(* Logix 5000 project; controller PLC_MCC1300_75F1 vendor 1 type 14 code 166 rev 32.11; software revision 32.04; part 13 of 83 *)
(* tags used below, declared in another part *)
   M302SpeedUp : MAC_SpeedUp;
   TMP_d : DINT;
   TMP_xPositioning : BOOL;
   TMP_xReverse : BOOL;
   TMP_xRun : BOOL;
   xAlwaysOFF : BOOL;
   Z300_Conveyor : UDT_StandConv[29];
   Z300_Conveyor_Conf : UDT_Conveyor_Config[29];
   Z300_Conveyor_HMW : MAC_Conveyor_ZC_HMW[29];
   Z300_Conveyor_IN_MOTION : MAC_Conveyor_ZC_IN_MOTION[29];
   Z301_HMR : MAC_Zone_ML_HMR;
(* CommandLogic, continued *)

ROUTINE M302M5_Conveyor_Output   (* ladder *)
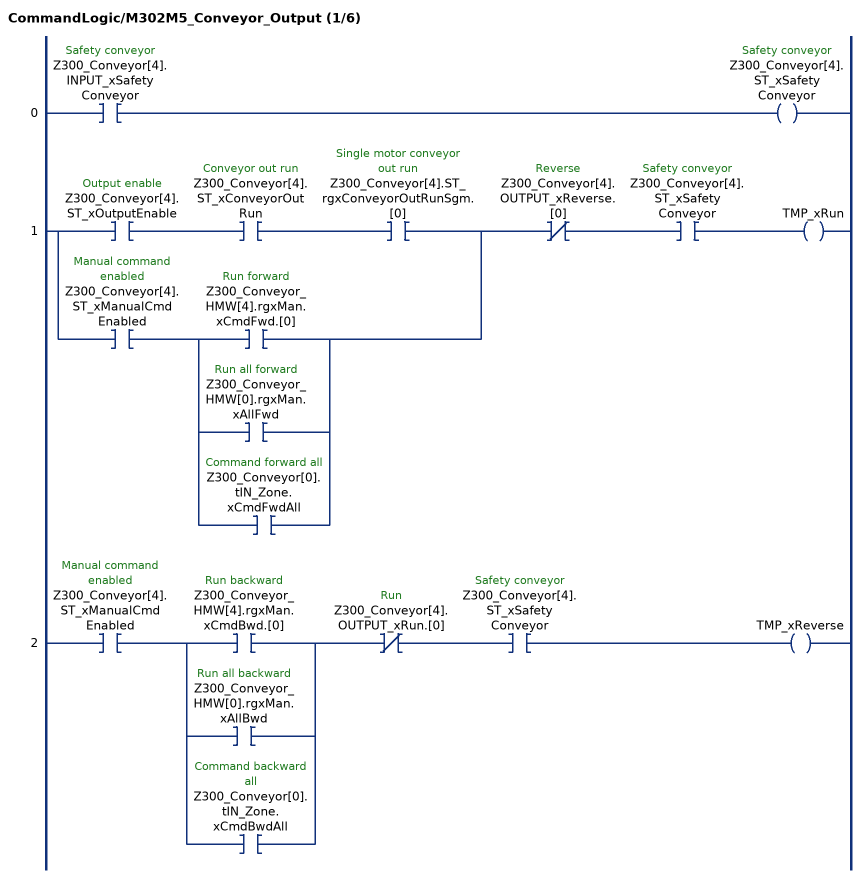
   0: XIC(Z300_Conveyor[4].INPUT_xSafetyConveyor)OTE(Z300_Conveyor[4].ST_xSafetyConveyor);
   1: [XIC(Z300_Conveyor[4].ST_xOutputEnable) XIC(Z300_Conveyor[4].ST_xConveyorOutRun) XIC(Z300_Conveyor[4].ST_rgxConveyorOutRunSgm.[0]) ,XIC(Z300_Conveyor[4].ST_xManualCmdEnabled) [XIC(Z300_Conveyor_HMW[4].rgxMan.xCmdFwd.[0]) ,XIC(Z300_Conveyor_HMW[0].rgxMan.xAllFwd) ,XIC(Z300_Conveyor[0].tIN_Zone.xCmdFwdAll) ] ]XIO(Z300_Conveyor[4].OUTPUT_xReverse.[0])XIC(Z300_Conveyor[4].ST_xSafetyConveyor)OTE(TMP_xRun);
   2: XIC(Z300_Conveyor[4].ST_xManualCmdEnabled)[XIC(Z300_Conveyor_HMW[4].rgxMan.xCmdBwd.[0]) ,XIC(Z300_Conveyor_HMW[0].rgxMan.xAllBwd) ,XIC(Z300_Conveyor[0].tIN_Zone.xCmdBwdAll) ]XIO(Z300_Conveyor[4].OUTPUT_xRun.[0])XIC(Z300_Conveyor[4].ST_xSafetyConveyor)OTE(TMP_xReverse);
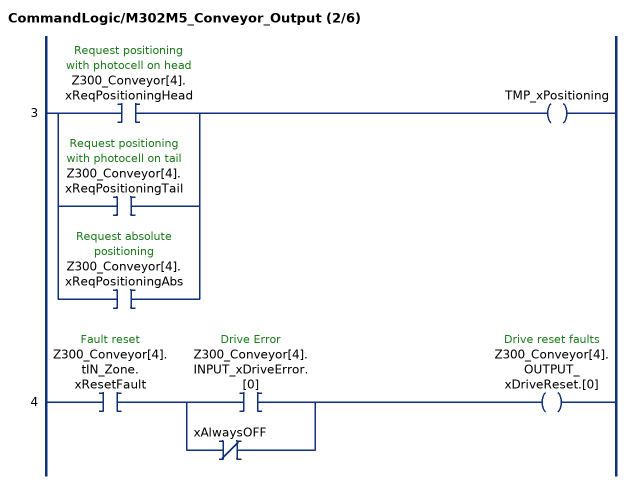
   3: [XIC(Z300_Conveyor[4].xReqPositioningHead) ,XIC(Z300_Conveyor[4].xReqPositioningTail) ,XIC(Z300_Conveyor[4].xReqPositioningAbs) ]OTE(TMP_xPositioning);
   4: XIC(Z300_Conveyor[4].tIN_Zone.xResetFault)[XIC(Z300_Conveyor[4].INPUT_xDriveError.[0]) ,XIO(xAlwaysOFF) ]OTE(Z300_Conveyor[4].OUTPUT_xDriveReset.[0]);
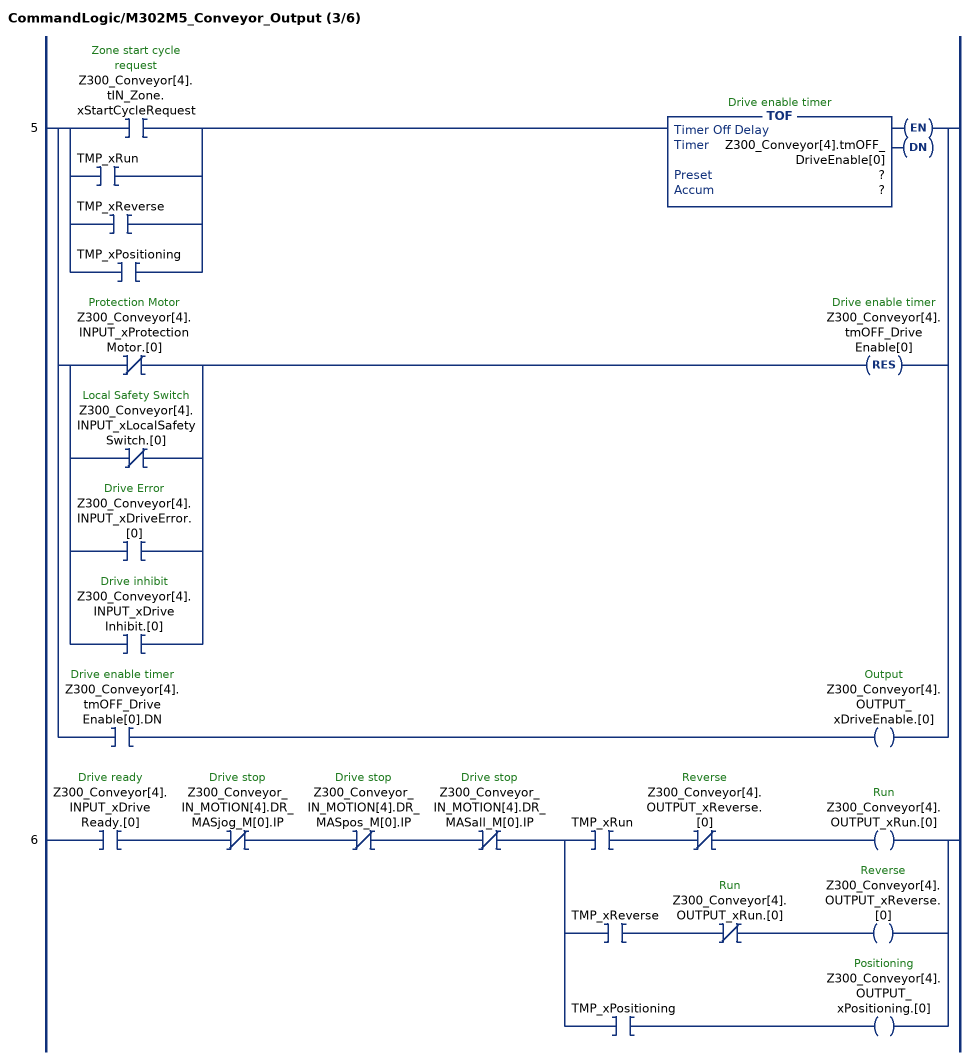
   5: [[XIC(Z300_Conveyor[4].tIN_Zone.xStartCycleRequest) ,XIC(TMP_xRun) ,XIC(TMP_xReverse) ,XIC(TMP_xPositioning) ] TOF(Z300_Conveyor[4].tmOFF_DriveEnable[0],?,?) ,[XIO(Z300_Conveyor[4].INPUT_xProtectionMotor.[0]) ,XIO(Z300_Conveyor[4].INPUT_xLocalSafetySwitch.[0]) ,XIC(Z300_Conveyor[4].INPUT_xDriveError.[0]) ,XIC(Z300_Conveyor[4].INPUT_xDriveInhibit.[0]) ] RES(Z300_Conveyor[4].tmOFF_DriveEnable[0]) ,XIC(Z300_Conveyor[4].tmOFF_DriveEnable[0].DN) OTE(Z300_Conveyor[4].OUTPUT_xDriveEnable.[0]) ];
   6: XIC(Z300_Conveyor[4].INPUT_xDriveReady.[0])XIO(Z300_Conveyor_IN_MOTION[4].DR_MASjog_M[0].IP)XIO(Z300_Conveyor_IN_MOTION[4].DR_MASpos_M[0].IP)XIO(Z300_Conveyor_IN_MOTION[4].DR_MASall_M[0].IP)[XIC(TMP_xRun) XIO(Z300_Conveyor[4].OUTPUT_xReverse.[0]) OTE(Z300_Conveyor[4].OUTPUT_xRun.[0]) ,XIC(TMP_xReverse) XIO(Z300_Conveyor[4].OUTPUT_xRun.[0]) OTE(Z300_Conveyor[4].OUTPUT_xReverse.[0]) ,XIC(TMP_xPositioning) OTE(Z300_Conveyor[4].OUTPUT_xPositioning.[0]) ];
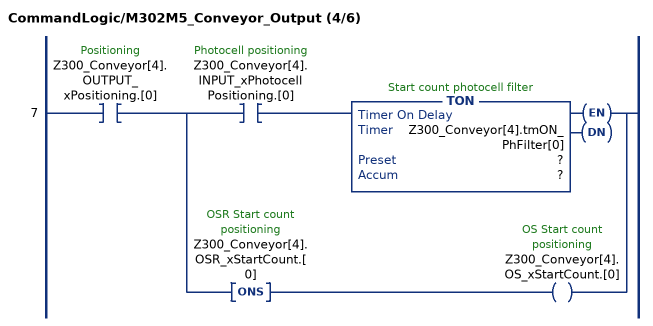
   7: XIC(Z300_Conveyor[4].OUTPUT_xPositioning.[0])[XIC(Z300_Conveyor[4].INPUT_xPhotocellPositioning.[0]) TON(Z300_Conveyor[4].tmON_PhFilter[0],?,?) ,ONS(Z300_Conveyor[4].OSR_xStartCount.[0]) OTE(Z300_Conveyor[4].OS_xStartCount.[0]) ];
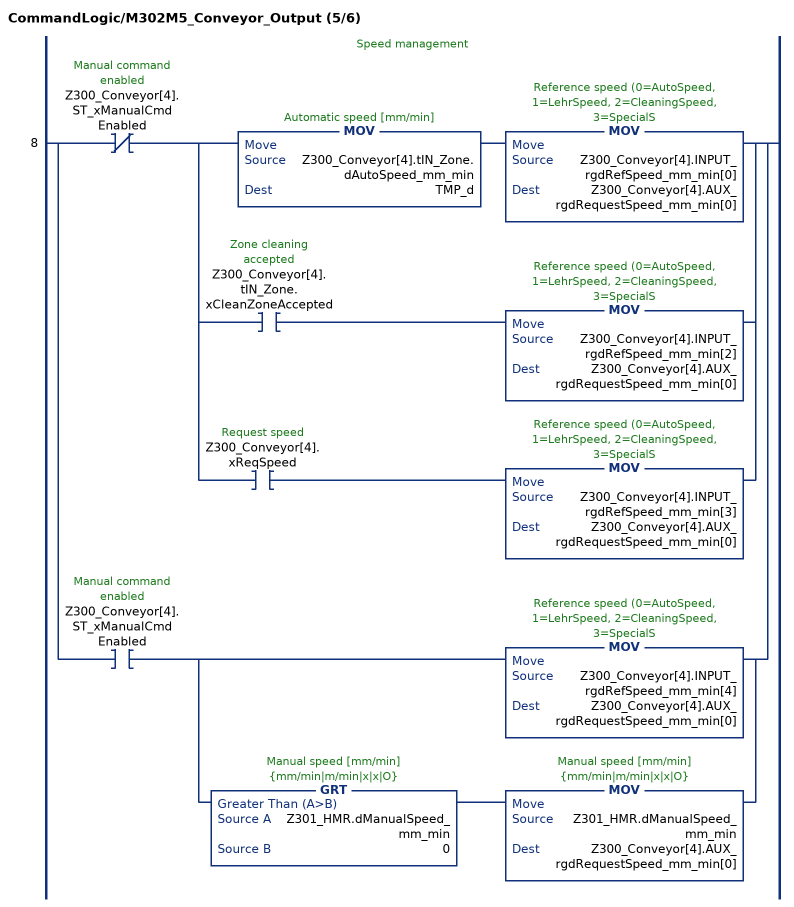
   // Speed management
   8: [XIO(Z300_Conveyor[4].ST_xManualCmdEnabled) [MOV(Z300_Conveyor[4].tIN_Zone.dAutoSpeed_mm_min,TMP_d) MOV(Z300_Conveyor[4].INPUT_rgdRefSpeed_mm_min[0],Z300_Conveyor[4].AUX_rgdRequestSpeed_mm_min[0]) ,XIC(Z300_Conveyor[4].tIN_Zone.xCleanZoneAccepted) MOV(Z300_Conveyor[4].INPUT_rgdRefSpeed_mm_min[2],Z300_Conveyor[4].AUX_rgdRequestSpeed_mm_min[0]) ,XIC(Z300_Conveyor[4].xReqSpeed) MOV(Z300_Conveyor[4].INPUT_rgdRefSpeed_mm_min[3],Z300_Conveyor[4].AUX_rgdRequestSpeed_mm_min[0]) ] ,XIC(Z300_Conveyor[4].ST_xManualCmdEnabled) [MOV(Z300_Conveyor[4].INPUT_rgdRefSpeed_mm_min[4],Z300_Conveyor[4].AUX_rgdRequestSpeed_mm_min[0]) ,GRT(Z301_HMR.dManualSpeed_mm_min,0) MOV(Z301_HMR.dManualSpeed_mm_min,Z300_Conveyor[4].AUX_rgdRequestSpeed_mm_min[0]) ] ];
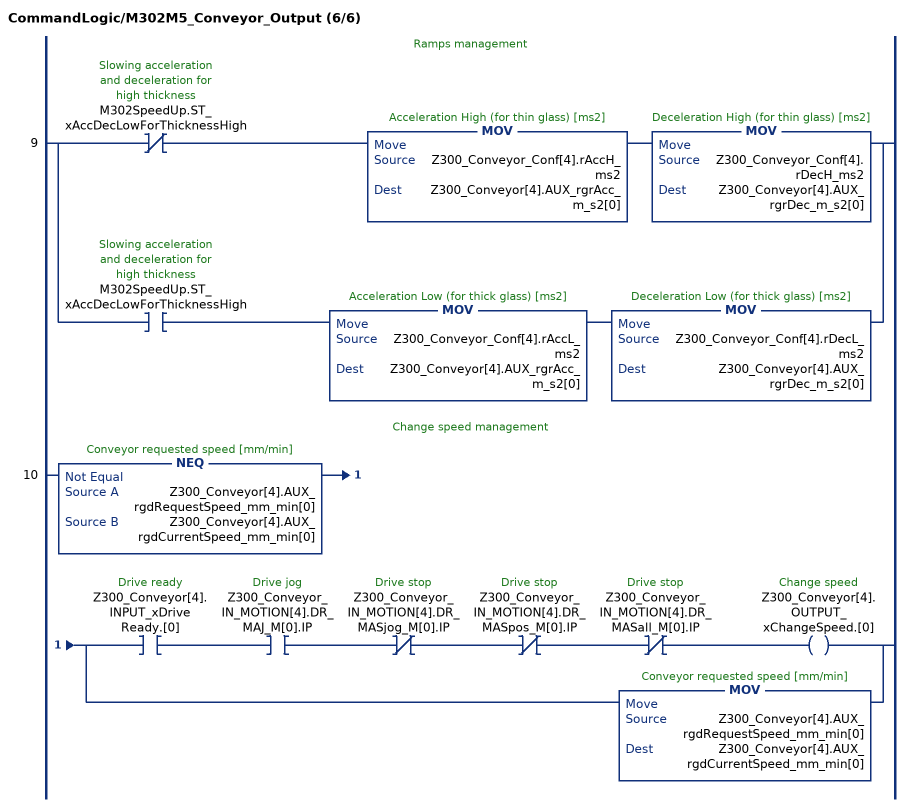
   // Ramps management
   9: [XIO(M302SpeedUp.ST_xAccDecLowForThicknessHigh) MOV(Z300_Conveyor_Conf[4].rAccH_ms2,Z300_Conveyor[4].AUX_rgrAcc_m_s2[0]) MOV(Z300_Conveyor_Conf[4].rDecH_ms2,Z300_Conveyor[4].AUX_rgrDec_m_s2[0]) ,XIC(M302SpeedUp.ST_xAccDecLowForThicknessHigh) MOV(Z300_Conveyor_Conf[4].rAccL_ms2,Z300_Conveyor[4].AUX_rgrAcc_m_s2[0]) MOV(Z300_Conveyor_Conf[4].rDecL_ms2,Z300_Conveyor[4].AUX_rgrDec_m_s2[0]) ];
   // Change speed management
   10: NEQ(Z300_Conveyor[4].AUX_rgdRequestSpeed_mm_min[0],Z300_Conveyor[4].AUX_rgdCurrentSpeed_mm_min[0])[XIC(Z300_Conveyor[4].INPUT_xDriveReady.[0]) XIC(Z300_Conveyor_IN_MOTION[4].DR_MAJ_M[0].IP) XIO(Z300_Conveyor_IN_MOTION[4].DR_MASjog_M[0].IP) XIO(Z300_Conveyor_IN_MOTION[4].DR_MASpos_M[0].IP) XIO(Z300_Conveyor_IN_MOTION[4].DR_MASall_M[0].IP) OTE(Z300_Conveyor[4].OUTPUT_xChangeSpeed.[0]) ,MOV(Z300_Conveyor[4].AUX_rgdRequestSpeed_mm_min[0],Z300_Conveyor[4].AUX_rgdCurrentSpeed_mm_min[0]) ];
END_ROUTINE

ROUTINE M302M6_Conveyor_Output   (* ladder *)
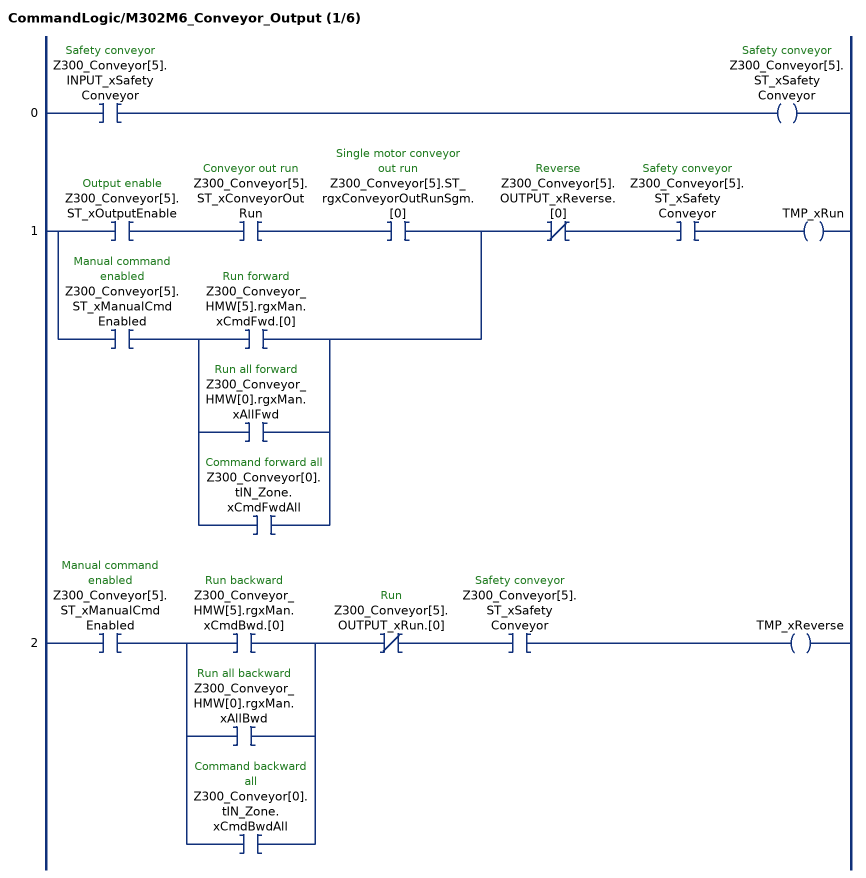
   0: XIC(Z300_Conveyor[5].INPUT_xSafetyConveyor)OTE(Z300_Conveyor[5].ST_xSafetyConveyor);
   1: [XIC(Z300_Conveyor[5].ST_xOutputEnable) XIC(Z300_Conveyor[5].ST_xConveyorOutRun) XIC(Z300_Conveyor[5].ST_rgxConveyorOutRunSgm.[0]) ,XIC(Z300_Conveyor[5].ST_xManualCmdEnabled) [XIC(Z300_Conveyor_HMW[5].rgxMan.xCmdFwd.[0]) ,XIC(Z300_Conveyor_HMW[0].rgxMan.xAllFwd) ,XIC(Z300_Conveyor[0].tIN_Zone.xCmdFwdAll) ] ]XIO(Z300_Conveyor[5].OUTPUT_xReverse.[0])XIC(Z300_Conveyor[5].ST_xSafetyConveyor)OTE(TMP_xRun);
   2: XIC(Z300_Conveyor[5].ST_xManualCmdEnabled)[XIC(Z300_Conveyor_HMW[5].rgxMan.xCmdBwd.[0]) ,XIC(Z300_Conveyor_HMW[0].rgxMan.xAllBwd) ,XIC(Z300_Conveyor[0].tIN_Zone.xCmdBwdAll) ]XIO(Z300_Conveyor[5].OUTPUT_xRun.[0])XIC(Z300_Conveyor[5].ST_xSafetyConveyor)OTE(TMP_xReverse);
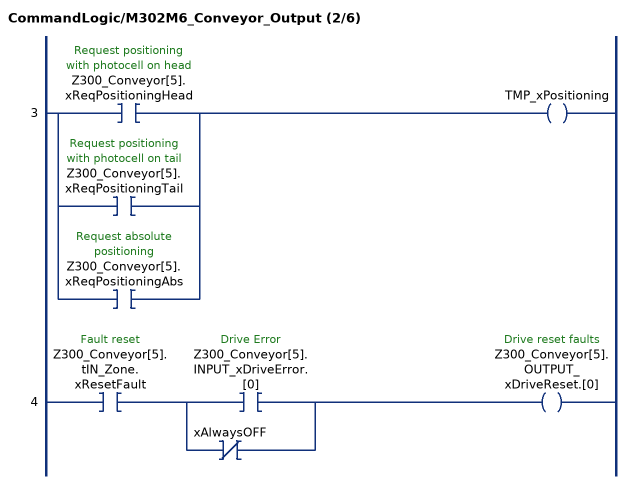
   3: [XIC(Z300_Conveyor[5].xReqPositioningHead) ,XIC(Z300_Conveyor[5].xReqPositioningTail) ,XIC(Z300_Conveyor[5].xReqPositioningAbs) ]OTE(TMP_xPositioning);
   4: XIC(Z300_Conveyor[5].tIN_Zone.xResetFault)[XIC(Z300_Conveyor[5].INPUT_xDriveError.[0]) ,XIO(xAlwaysOFF) ]OTE(Z300_Conveyor[5].OUTPUT_xDriveReset.[0]);
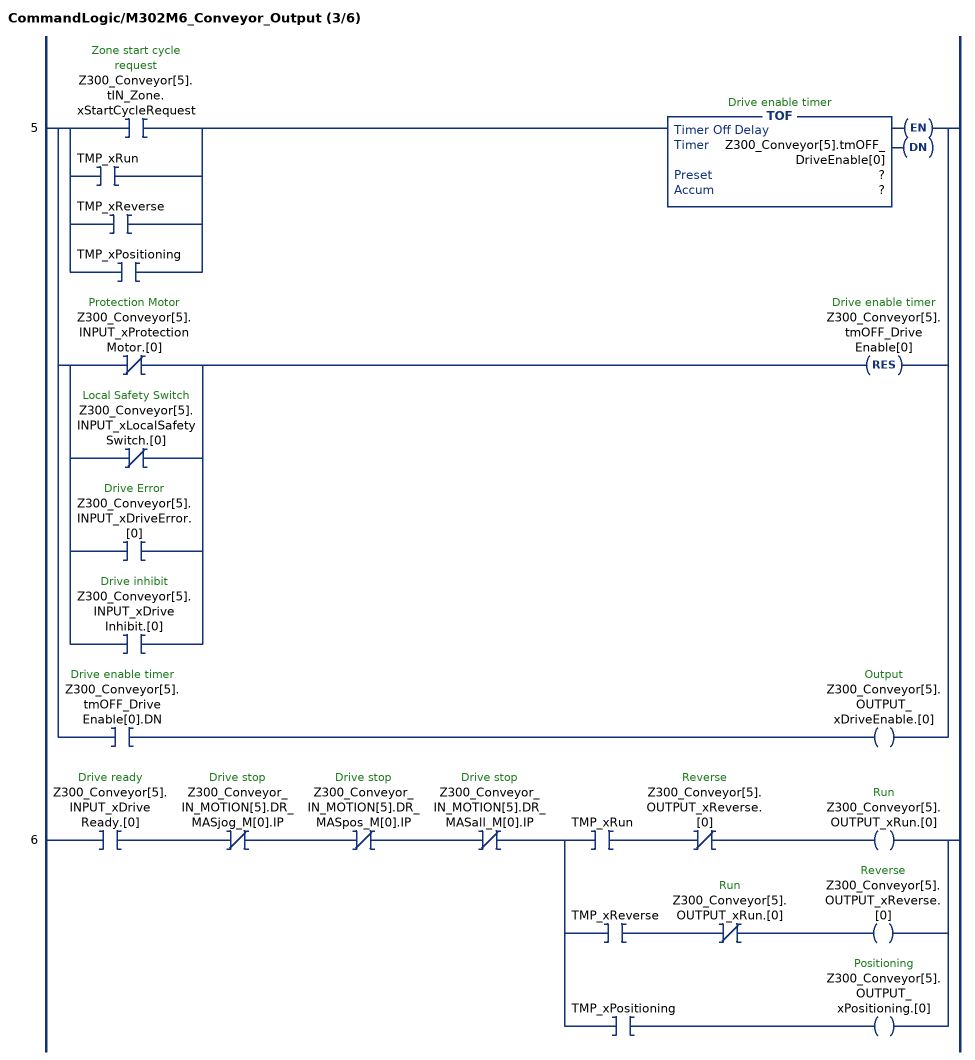
   5: [[XIC(Z300_Conveyor[5].tIN_Zone.xStartCycleRequest) ,XIC(TMP_xRun) ,XIC(TMP_xReverse) ,XIC(TMP_xPositioning) ] TOF(Z300_Conveyor[5].tmOFF_DriveEnable[0],?,?) ,[XIO(Z300_Conveyor[5].INPUT_xProtectionMotor.[0]) ,XIO(Z300_Conveyor[5].INPUT_xLocalSafetySwitch.[0]) ,XIC(Z300_Conveyor[5].INPUT_xDriveError.[0]) ,XIC(Z300_Conveyor[5].INPUT_xDriveInhibit.[0]) ] RES(Z300_Conveyor[5].tmOFF_DriveEnable[0]) ,XIC(Z300_Conveyor[5].tmOFF_DriveEnable[0].DN) OTE(Z300_Conveyor[5].OUTPUT_xDriveEnable.[0]) ];
   6: XIC(Z300_Conveyor[5].INPUT_xDriveReady.[0])XIO(Z300_Conveyor_IN_MOTION[5].DR_MASjog_M[0].IP)XIO(Z300_Conveyor_IN_MOTION[5].DR_MASpos_M[0].IP)XIO(Z300_Conveyor_IN_MOTION[5].DR_MASall_M[0].IP)[XIC(TMP_xRun) XIO(Z300_Conveyor[5].OUTPUT_xReverse.[0]) OTE(Z300_Conveyor[5].OUTPUT_xRun.[0]) ,XIC(TMP_xReverse) XIO(Z300_Conveyor[5].OUTPUT_xRun.[0]) OTE(Z300_Conveyor[5].OUTPUT_xReverse.[0]) ,XIC(TMP_xPositioning) OTE(Z300_Conveyor[5].OUTPUT_xPositioning.[0]) ];
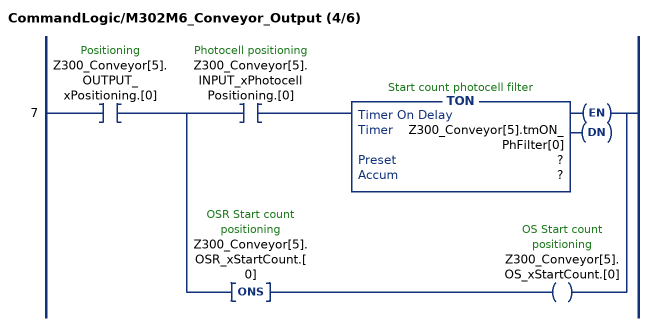
   7: XIC(Z300_Conveyor[5].OUTPUT_xPositioning.[0])[XIC(Z300_Conveyor[5].INPUT_xPhotocellPositioning.[0]) TON(Z300_Conveyor[5].tmON_PhFilter[0],?,?) ,ONS(Z300_Conveyor[5].OSR_xStartCount.[0]) OTE(Z300_Conveyor[5].OS_xStartCount.[0]) ];
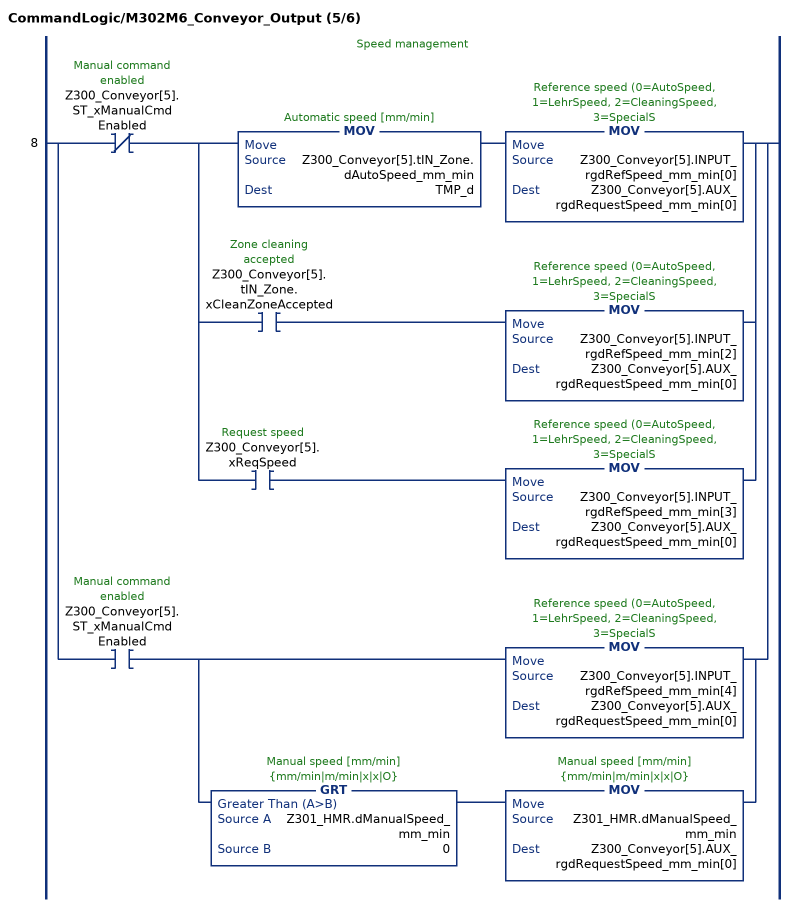
   // Speed management
   8: [XIO(Z300_Conveyor[5].ST_xManualCmdEnabled) [MOV(Z300_Conveyor[5].tIN_Zone.dAutoSpeed_mm_min,TMP_d) MOV(Z300_Conveyor[5].INPUT_rgdRefSpeed_mm_min[0],Z300_Conveyor[5].AUX_rgdRequestSpeed_mm_min[0]) ,XIC(Z300_Conveyor[5].tIN_Zone.xCleanZoneAccepted) MOV(Z300_Conveyor[5].INPUT_rgdRefSpeed_mm_min[2],Z300_Conveyor[5].AUX_rgdRequestSpeed_mm_min[0]) ,XIC(Z300_Conveyor[5].xReqSpeed) MOV(Z300_Conveyor[5].INPUT_rgdRefSpeed_mm_min[3],Z300_Conveyor[5].AUX_rgdRequestSpeed_mm_min[0]) ] ,XIC(Z300_Conveyor[5].ST_xManualCmdEnabled) [MOV(Z300_Conveyor[5].INPUT_rgdRefSpeed_mm_min[4],Z300_Conveyor[5].AUX_rgdRequestSpeed_mm_min[0]) ,GRT(Z301_HMR.dManualSpeed_mm_min,0) MOV(Z301_HMR.dManualSpeed_mm_min,Z300_Conveyor[5].AUX_rgdRequestSpeed_mm_min[0]) ] ];
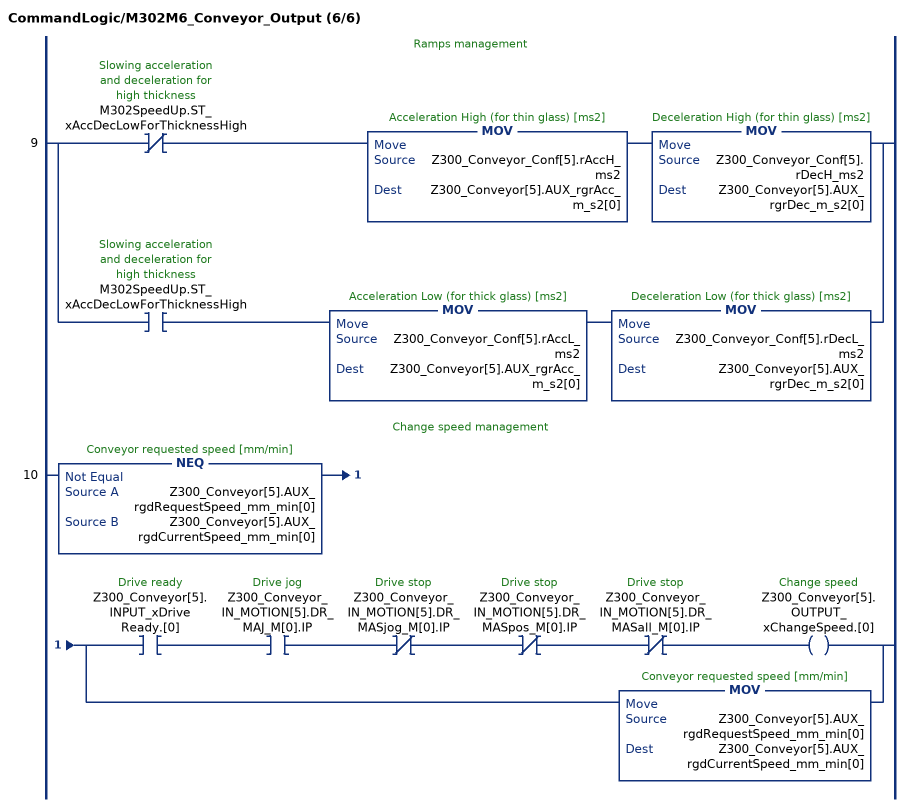
   // Ramps management
   9: [XIO(M302SpeedUp.ST_xAccDecLowForThicknessHigh) MOV(Z300_Conveyor_Conf[5].rAccH_ms2,Z300_Conveyor[5].AUX_rgrAcc_m_s2[0]) MOV(Z300_Conveyor_Conf[5].rDecH_ms2,Z300_Conveyor[5].AUX_rgrDec_m_s2[0]) ,XIC(M302SpeedUp.ST_xAccDecLowForThicknessHigh) MOV(Z300_Conveyor_Conf[5].rAccL_ms2,Z300_Conveyor[5].AUX_rgrAcc_m_s2[0]) MOV(Z300_Conveyor_Conf[5].rDecL_ms2,Z300_Conveyor[5].AUX_rgrDec_m_s2[0]) ];
   // Change speed management
   10: NEQ(Z300_Conveyor[5].AUX_rgdRequestSpeed_mm_min[0],Z300_Conveyor[5].AUX_rgdCurrentSpeed_mm_min[0])[XIC(Z300_Conveyor[5].INPUT_xDriveReady.[0]) XIC(Z300_Conveyor_IN_MOTION[5].DR_MAJ_M[0].IP) XIO(Z300_Conveyor_IN_MOTION[5].DR_MASjog_M[0].IP) XIO(Z300_Conveyor_IN_MOTION[5].DR_MASpos_M[0].IP) XIO(Z300_Conveyor_IN_MOTION[5].DR_MASall_M[0].IP) OTE(Z300_Conveyor[5].OUTPUT_xChangeSpeed.[0]) ,MOV(Z300_Conveyor[5].AUX_rgdRequestSpeed_mm_min[0],Z300_Conveyor[5].AUX_rgdCurrentSpeed_mm_min[0]) ];
END_ROUTINE

ROUTINE M302M7_Conveyor_Output   (* ladder *)
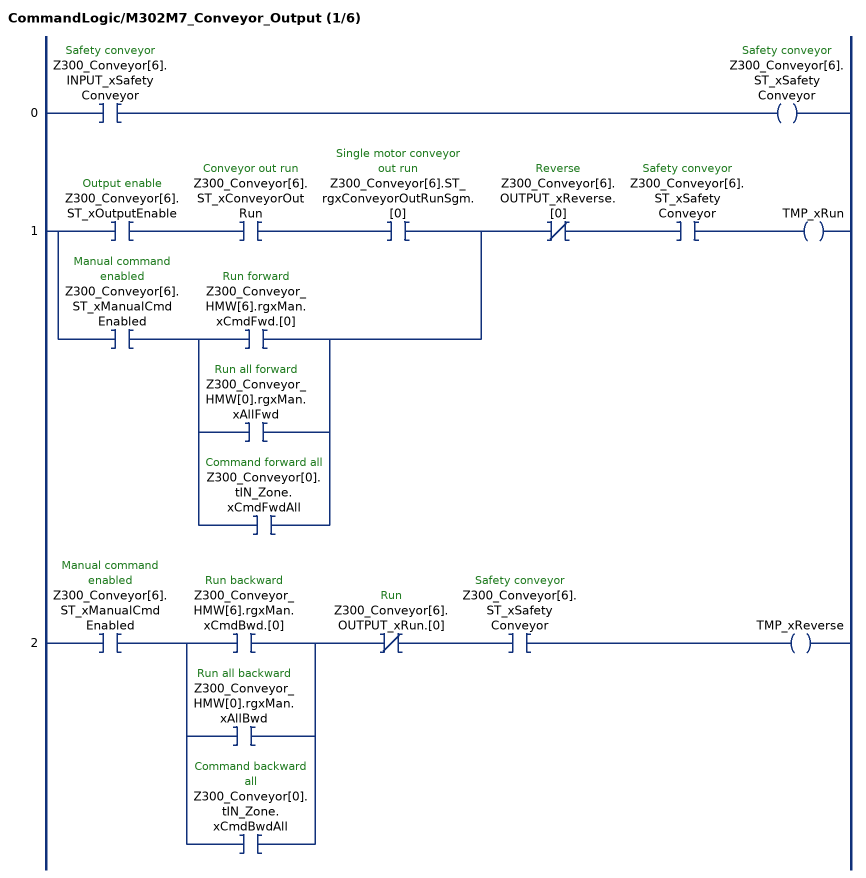
   0: XIC(Z300_Conveyor[6].INPUT_xSafetyConveyor)OTE(Z300_Conveyor[6].ST_xSafetyConveyor);
   1: [XIC(Z300_Conveyor[6].ST_xOutputEnable) XIC(Z300_Conveyor[6].ST_xConveyorOutRun) XIC(Z300_Conveyor[6].ST_rgxConveyorOutRunSgm.[0]) ,XIC(Z300_Conveyor[6].ST_xManualCmdEnabled) [XIC(Z300_Conveyor_HMW[6].rgxMan.xCmdFwd.[0]) ,XIC(Z300_Conveyor_HMW[0].rgxMan.xAllFwd) ,XIC(Z300_Conveyor[0].tIN_Zone.xCmdFwdAll) ] ]XIO(Z300_Conveyor[6].OUTPUT_xReverse.[0])XIC(Z300_Conveyor[6].ST_xSafetyConveyor)OTE(TMP_xRun);
   2: XIC(Z300_Conveyor[6].ST_xManualCmdEnabled)[XIC(Z300_Conveyor_HMW[6].rgxMan.xCmdBwd.[0]) ,XIC(Z300_Conveyor_HMW[0].rgxMan.xAllBwd) ,XIC(Z300_Conveyor[0].tIN_Zone.xCmdBwdAll) ]XIO(Z300_Conveyor[6].OUTPUT_xRun.[0])XIC(Z300_Conveyor[6].ST_xSafetyConveyor)OTE(TMP_xReverse);
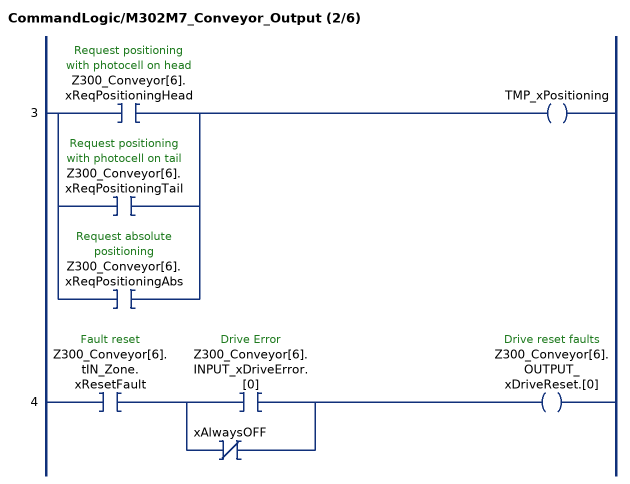
   3: [XIC(Z300_Conveyor[6].xReqPositioningHead) ,XIC(Z300_Conveyor[6].xReqPositioningTail) ,XIC(Z300_Conveyor[6].xReqPositioningAbs) ]OTE(TMP_xPositioning);
   4: XIC(Z300_Conveyor[6].tIN_Zone.xResetFault)[XIC(Z300_Conveyor[6].INPUT_xDriveError.[0]) ,XIO(xAlwaysOFF) ]OTE(Z300_Conveyor[6].OUTPUT_xDriveReset.[0]);
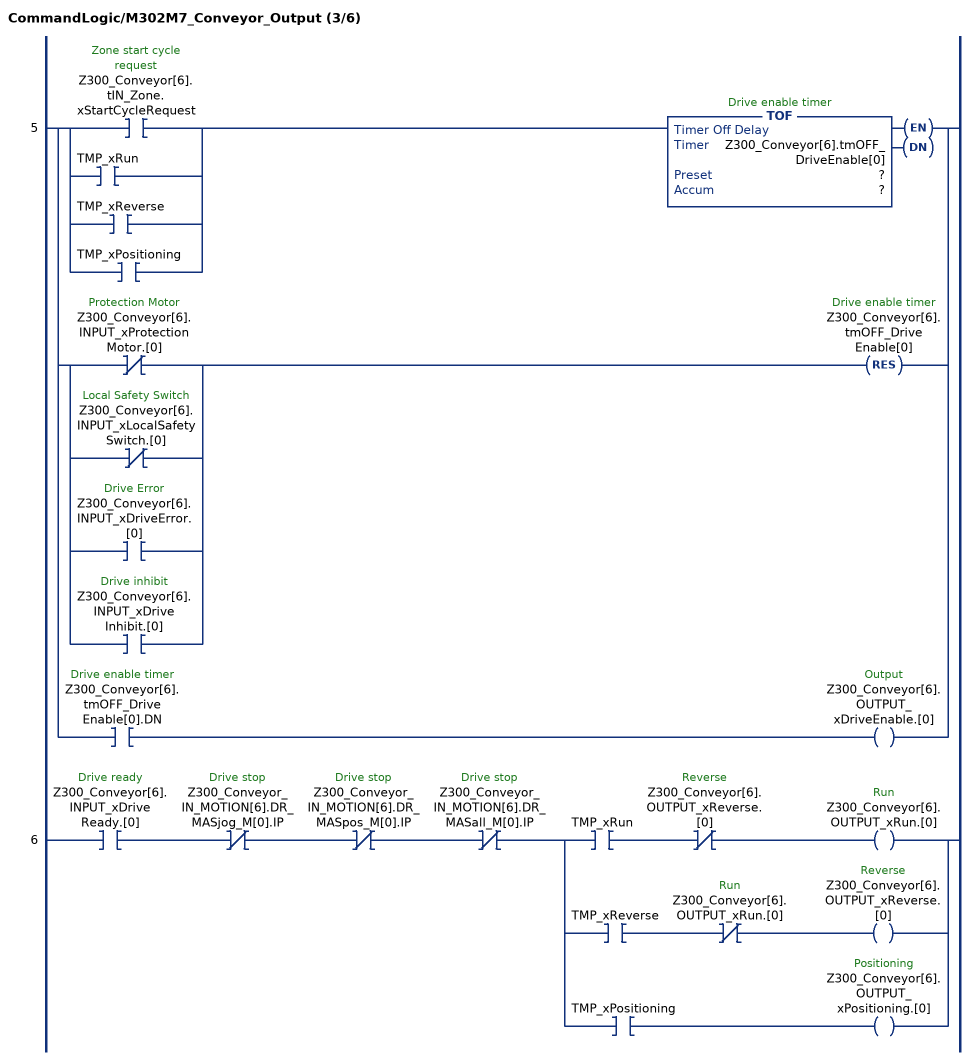
   5: [[XIC(Z300_Conveyor[6].tIN_Zone.xStartCycleRequest) ,XIC(TMP_xRun) ,XIC(TMP_xReverse) ,XIC(TMP_xPositioning) ] TOF(Z300_Conveyor[6].tmOFF_DriveEnable[0],?,?) ,[XIO(Z300_Conveyor[6].INPUT_xProtectionMotor.[0]) ,XIO(Z300_Conveyor[6].INPUT_xLocalSafetySwitch.[0]) ,XIC(Z300_Conveyor[6].INPUT_xDriveError.[0]) ,XIC(Z300_Conveyor[6].INPUT_xDriveInhibit.[0]) ] RES(Z300_Conveyor[6].tmOFF_DriveEnable[0]) ,XIC(Z300_Conveyor[6].tmOFF_DriveEnable[0].DN) OTE(Z300_Conveyor[6].OUTPUT_xDriveEnable.[0]) ];
   6: XIC(Z300_Conveyor[6].INPUT_xDriveReady.[0])XIO(Z300_Conveyor_IN_MOTION[6].DR_MASjog_M[0].IP)XIO(Z300_Conveyor_IN_MOTION[6].DR_MASpos_M[0].IP)XIO(Z300_Conveyor_IN_MOTION[6].DR_MASall_M[0].IP)[XIC(TMP_xRun) XIO(Z300_Conveyor[6].OUTPUT_xReverse.[0]) OTE(Z300_Conveyor[6].OUTPUT_xRun.[0]) ,XIC(TMP_xReverse) XIO(Z300_Conveyor[6].OUTPUT_xRun.[0]) OTE(Z300_Conveyor[6].OUTPUT_xReverse.[0]) ,XIC(TMP_xPositioning) OTE(Z300_Conveyor[6].OUTPUT_xPositioning.[0]) ];
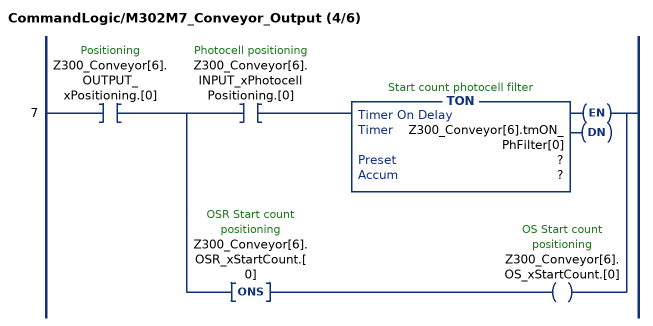
   7: XIC(Z300_Conveyor[6].OUTPUT_xPositioning.[0])[XIC(Z300_Conveyor[6].INPUT_xPhotocellPositioning.[0]) TON(Z300_Conveyor[6].tmON_PhFilter[0],?,?) ,ONS(Z300_Conveyor[6].OSR_xStartCount.[0]) OTE(Z300_Conveyor[6].OS_xStartCount.[0]) ];
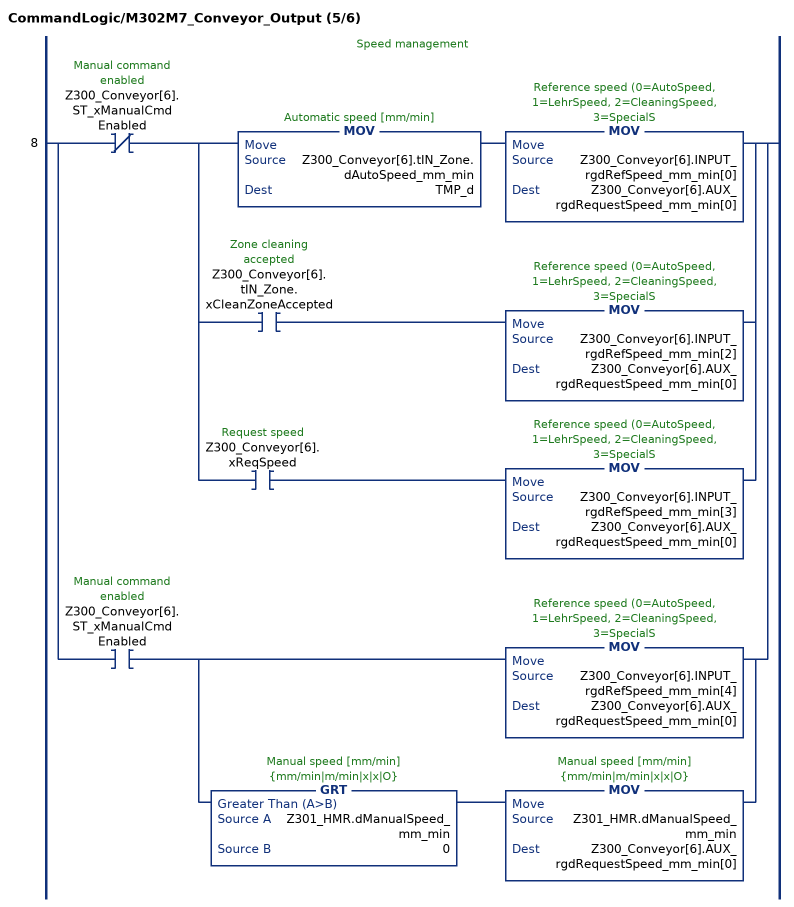
   // Speed management
   8: [XIO(Z300_Conveyor[6].ST_xManualCmdEnabled) [MOV(Z300_Conveyor[6].tIN_Zone.dAutoSpeed_mm_min,TMP_d) MOV(Z300_Conveyor[6].INPUT_rgdRefSpeed_mm_min[0],Z300_Conveyor[6].AUX_rgdRequestSpeed_mm_min[0]) ,XIC(Z300_Conveyor[6].tIN_Zone.xCleanZoneAccepted) MOV(Z300_Conveyor[6].INPUT_rgdRefSpeed_mm_min[2],Z300_Conveyor[6].AUX_rgdRequestSpeed_mm_min[0]) ,XIC(Z300_Conveyor[6].xReqSpeed) MOV(Z300_Conveyor[6].INPUT_rgdRefSpeed_mm_min[3],Z300_Conveyor[6].AUX_rgdRequestSpeed_mm_min[0]) ] ,XIC(Z300_Conveyor[6].ST_xManualCmdEnabled) [MOV(Z300_Conveyor[6].INPUT_rgdRefSpeed_mm_min[4],Z300_Conveyor[6].AUX_rgdRequestSpeed_mm_min[0]) ,GRT(Z301_HMR.dManualSpeed_mm_min,0) MOV(Z301_HMR.dManualSpeed_mm_min,Z300_Conveyor[6].AUX_rgdRequestSpeed_mm_min[0]) ] ];
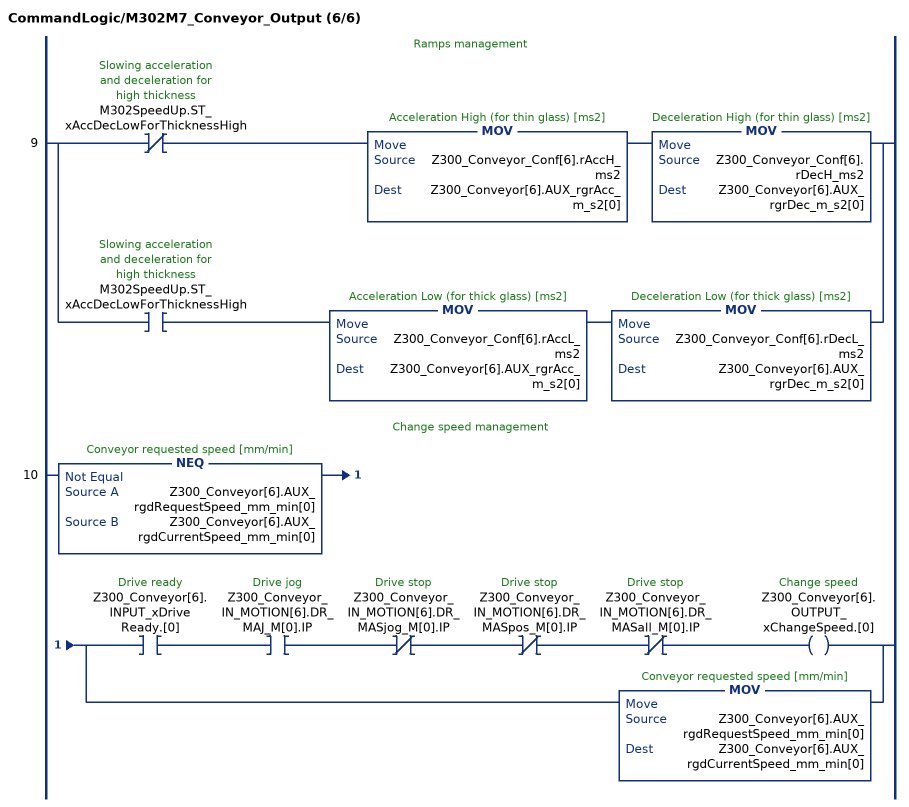
   // Ramps management
   9: [XIO(M302SpeedUp.ST_xAccDecLowForThicknessHigh) MOV(Z300_Conveyor_Conf[6].rAccH_ms2,Z300_Conveyor[6].AUX_rgrAcc_m_s2[0]) MOV(Z300_Conveyor_Conf[6].rDecH_ms2,Z300_Conveyor[6].AUX_rgrDec_m_s2[0]) ,XIC(M302SpeedUp.ST_xAccDecLowForThicknessHigh) MOV(Z300_Conveyor_Conf[6].rAccL_ms2,Z300_Conveyor[6].AUX_rgrAcc_m_s2[0]) MOV(Z300_Conveyor_Conf[6].rDecL_ms2,Z300_Conveyor[6].AUX_rgrDec_m_s2[0]) ];
   // Change speed management
   10: NEQ(Z300_Conveyor[6].AUX_rgdRequestSpeed_mm_min[0],Z300_Conveyor[6].AUX_rgdCurrentSpeed_mm_min[0])[XIC(Z300_Conveyor[6].INPUT_xDriveReady.[0]) XIC(Z300_Conveyor_IN_MOTION[6].DR_MAJ_M[0].IP) XIO(Z300_Conveyor_IN_MOTION[6].DR_MASjog_M[0].IP) XIO(Z300_Conveyor_IN_MOTION[6].DR_MASpos_M[0].IP) XIO(Z300_Conveyor_IN_MOTION[6].DR_MASall_M[0].IP) OTE(Z300_Conveyor[6].OUTPUT_xChangeSpeed.[0]) ,MOV(Z300_Conveyor[6].AUX_rgdRequestSpeed_mm_min[0],Z300_Conveyor[6].AUX_rgdCurrentSpeed_mm_min[0]) ];
END_ROUTINE
